REGION Network 319: CARRIER ENCODER POSITION FAULT
   RUNG wire#powerrail
      Contact( "reset" )
      { S7_Templates := "SrcType := Word" } EQ_Contact(in1 := "DB101_DB_SDC_FAULTS".Carrier_Fault[39], in2 := 131)
      Coil( "DB302_HMI_Faults".Carrier39_Faults_0.%X12 )
   END_RUNG
   // the same network as SCL:
   "DB302_HMI_Faults".Carrier39_Faults_0.%X12 := "reset" AND ("DB101_DB_SDC_FAULTS".Carrier_Fault[39] = 131);
END_REGION

REGION Network 320: CARRIER ENCODER INTERNAL ERROR
   RUNG wire#powerrail
      Contact( "reset" )
      { S7_Templates := "SrcType := Word" } EQ_Contact(in1 := "DB101_DB_SDC_FAULTS".Carrier_Fault[39], in2 := 132)
      Coil( "DB302_HMI_Faults".Carrier39_Faults_0.%X13 )
   END_RUNG
   // the same network as SCL:
   "DB302_HMI_Faults".Carrier39_Faults_0.%X13 := "reset" AND ("DB101_DB_SDC_FAULTS".Carrier_Fault[39] = 132);
END_REGION

REGION Network 321: CARRIER ENCODER COMM FAULT
   RUNG wire#powerrail
      Contact( "reset" )
      { S7_Templates := "SrcType := Word" } EQ_Contact(in1 := "DB101_DB_SDC_FAULTS".Carrier_Fault[39], in2 := 133)
      Coil( "DB302_HMI_Faults".Carrier39_Faults_0.%X14 )
   END_RUNG
   // the same network as SCL:
   "DB302_HMI_Faults".Carrier39_Faults_0.%X14 := "reset" AND ("DB101_DB_SDC_FAULTS".Carrier_Fault[39] = 133);
END_REGION

REGION Network 322: CARRIER HMI COMM FAULT
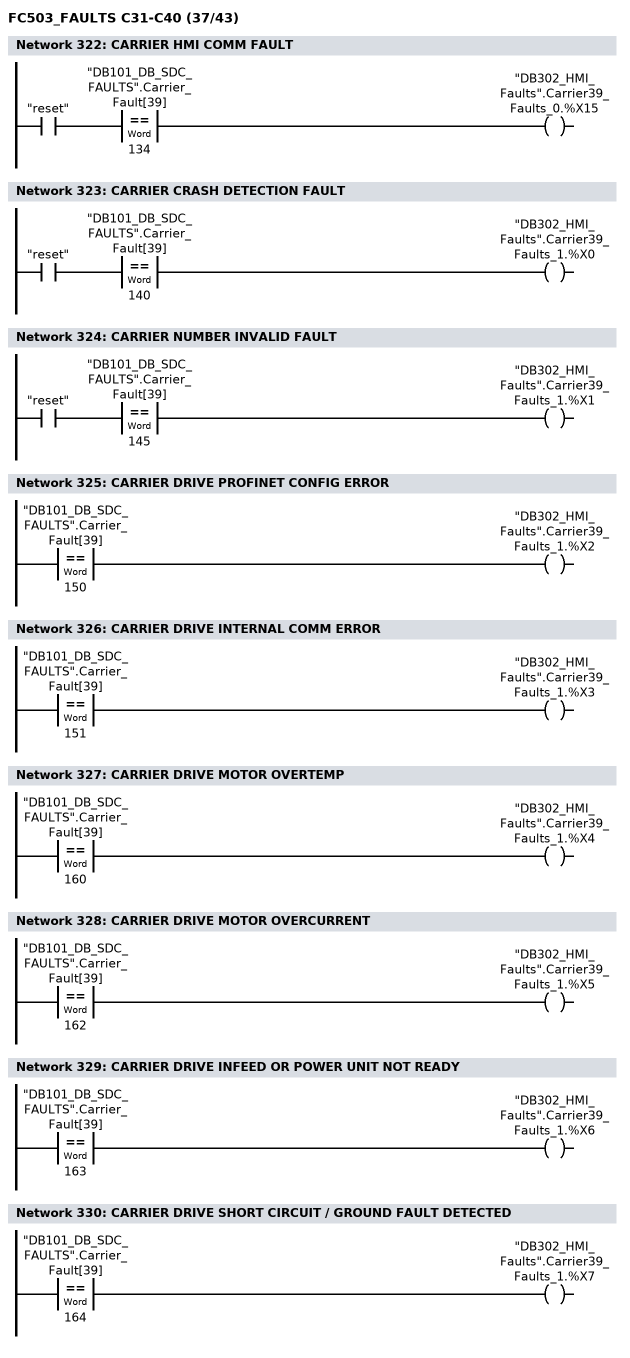
   RUNG wire#powerrail
      Contact( "reset" )
      { S7_Templates := "SrcType := Word" } EQ_Contact(in1 := "DB101_DB_SDC_FAULTS".Carrier_Fault[39], in2 := 134)
      Coil( "DB302_HMI_Faults".Carrier39_Faults_0.%X15 )
   END_RUNG
   // the same network as SCL:
   "DB302_HMI_Faults".Carrier39_Faults_0.%X15 := "reset" AND ("DB101_DB_SDC_FAULTS".Carrier_Fault[39] = 134);
END_REGION

REGION Network 323: CARRIER CRASH DETECTION FAULT
   RUNG wire#powerrail
      Contact( "reset" )
      { S7_Templates := "SrcType := Word" } EQ_Contact(in1 := "DB101_DB_SDC_FAULTS".Carrier_Fault[39], in2 := 140)
      Coil( "DB302_HMI_Faults".Carrier39_Faults_1.%X0 )
   END_RUNG
   // the same network as SCL:
   "DB302_HMI_Faults".Carrier39_Faults_1.%X0 := "reset" AND ("DB101_DB_SDC_FAULTS".Carrier_Fault[39] = 140);
END_REGION

REGION Network 324: CARRIER NUMBER INVALID FAULT
   RUNG wire#powerrail
      Contact( "reset" )
      { S7_Templates := "SrcType := Word" } EQ_Contact(in1 := "DB101_DB_SDC_FAULTS".Carrier_Fault[39], in2 := 145)
      Coil( "DB302_HMI_Faults".Carrier39_Faults_1.%X1 )
   END_RUNG
   // the same network as SCL:
   "DB302_HMI_Faults".Carrier39_Faults_1.%X1 := "reset" AND ("DB101_DB_SDC_FAULTS".Carrier_Fault[39] = 145);
END_REGION

REGION Network 325: CARRIER DRIVE PROFINET CONFIG ERROR
   RUNG wire#powerrail
      { S7_Templates := "SrcType := Word" } EQ_Contact(in1 := "DB101_DB_SDC_FAULTS".Carrier_Fault[39], in2 := 150)
      Coil( "DB302_HMI_Faults".Carrier39_Faults_1.%X2 )
   END_RUNG
   // the same network as SCL:
   "DB302_HMI_Faults".Carrier39_Faults_1.%X2 := "DB101_DB_SDC_FAULTS".Carrier_Fault[39] = 150;
END_REGION

REGION Network 326: CARRIER DRIVE INTERNAL COMM ERROR
   RUNG wire#powerrail
      { S7_Templates := "SrcType := Word" } EQ_Contact(in1 := "DB101_DB_SDC_FAULTS".Carrier_Fault[39], in2 := 151)
      Coil( "DB302_HMI_Faults".Carrier39_Faults_1.%X3 )
   END_RUNG
   // the same network as SCL:
   "DB302_HMI_Faults".Carrier39_Faults_1.%X3 := "DB101_DB_SDC_FAULTS".Carrier_Fault[39] = 151;
END_REGION

REGION Network 327: CARRIER DRIVE MOTOR OVERTEMP
   RUNG wire#powerrail
      { S7_Templates := "SrcType := Word" } EQ_Contact(in1 := "DB101_DB_SDC_FAULTS".Carrier_Fault[39], in2 := 160)
      Coil( "DB302_HMI_Faults".Carrier39_Faults_1.%X4 )
   END_RUNG
   // the same network as SCL:
   "DB302_HMI_Faults".Carrier39_Faults_1.%X4 := "DB101_DB_SDC_FAULTS".Carrier_Fault[39] = 160;
END_REGION

REGION Network 328: CARRIER DRIVE MOTOR OVERCURRENT
   RUNG wire#powerrail
      { S7_Templates := "SrcType := Word" } EQ_Contact(in1 := "DB101_DB_SDC_FAULTS".Carrier_Fault[39], in2 := 162)
      Coil( "DB302_HMI_Faults".Carrier39_Faults_1.%X5 )
   END_RUNG
   // the same network as SCL:
   "DB302_HMI_Faults".Carrier39_Faults_1.%X5 := "DB101_DB_SDC_FAULTS".Carrier_Fault[39] = 162;
END_REGION

REGION Network 329: CARRIER DRIVE INFEED OR POWER UNIT NOT READY
   RUNG wire#powerrail
      { S7_Templates := "SrcType := Word" } EQ_Contact(in1 := "DB101_DB_SDC_FAULTS".Carrier_Fault[39], in2 := 163)
      Coil( "DB302_HMI_Faults".Carrier39_Faults_1.%X6 )
   END_RUNG
   // the same network as SCL:
   "DB302_HMI_Faults".Carrier39_Faults_1.%X6 := "DB101_DB_SDC_FAULTS".Carrier_Fault[39] = 163;
END_REGION

REGION Network 330: CARRIER DRIVE SHORT CIRCUIT / GROUND FAULT DETECTED
   RUNG wire#powerrail
      { S7_Templates := "SrcType := Word" } EQ_Contact(in1 := "DB101_DB_SDC_FAULTS".Carrier_Fault[39], in2 := 164)
      Coil( "DB302_HMI_Faults".Carrier39_Faults_1.%X7 )
   END_RUNG
   // the same network as SCL:
   "DB302_HMI_Faults".Carrier39_Faults_1.%X7 := "DB101_DB_SDC_FAULTS".Carrier_Fault[39] = 164;
END_REGION

REGION Network 331: CARRIER DRIVE PROFINET SETPOINT TIMEOUT
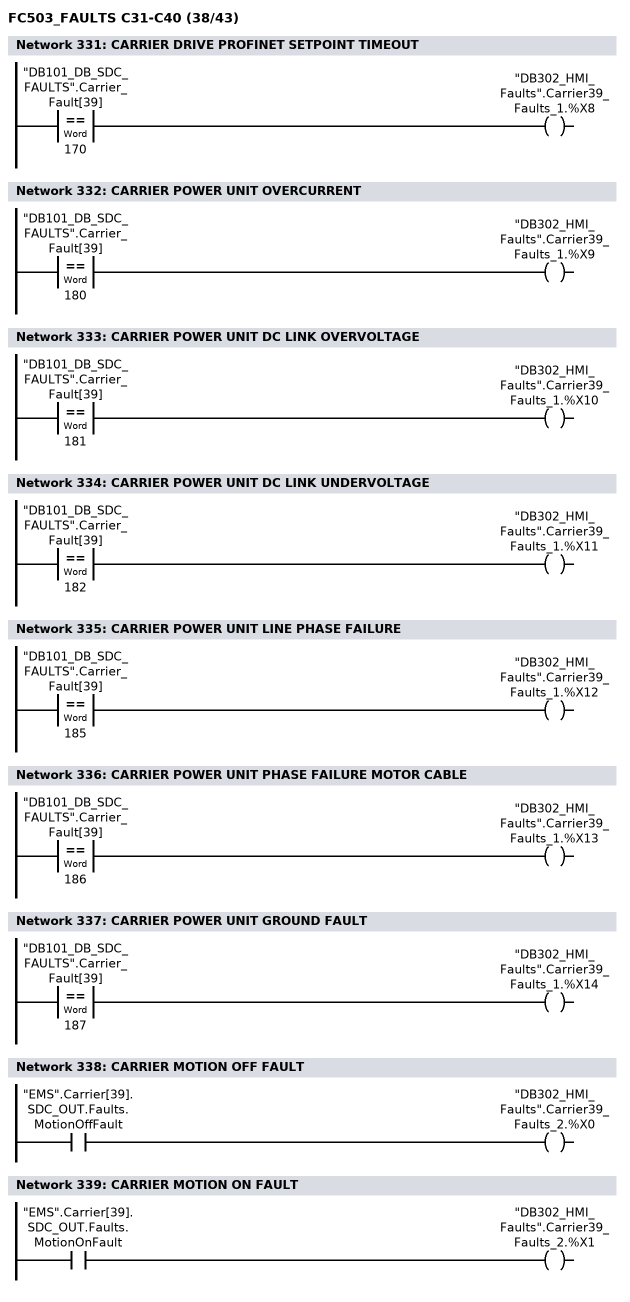
   RUNG wire#powerrail
      { S7_Templates := "SrcType := Word" } EQ_Contact(in1 := "DB101_DB_SDC_FAULTS".Carrier_Fault[39], in2 := 170)
      Coil( "DB302_HMI_Faults".Carrier39_Faults_1.%X8 )
   END_RUNG
   // the same network as SCL:
   "DB302_HMI_Faults".Carrier39_Faults_1.%X8 := "DB101_DB_SDC_FAULTS".Carrier_Fault[39] = 170;
END_REGION

REGION Network 332: CARRIER POWER UNIT OVERCURRENT
   RUNG wire#powerrail
      { S7_Templates := "SrcType := Word" } EQ_Contact(in1 := "DB101_DB_SDC_FAULTS".Carrier_Fault[39], in2 := 180)
      Coil( "DB302_HMI_Faults".Carrier39_Faults_1.%X9 )
   END_RUNG
   // the same network as SCL:
   "DB302_HMI_Faults".Carrier39_Faults_1.%X9 := "DB101_DB_SDC_FAULTS".Carrier_Fault[39] = 180;
END_REGION

REGION Network 333: CARRIER POWER UNIT DC LINK OVERVOLTAGE
   RUNG wire#powerrail
      { S7_Templates := "SrcType := Word" } EQ_Contact(in1 := "DB101_DB_SDC_FAULTS".Carrier_Fault[39], in2 := 181)
      Coil( "DB302_HMI_Faults".Carrier39_Faults_1.%X10 )
   END_RUNG
   // the same network as SCL:
   "DB302_HMI_Faults".Carrier39_Faults_1.%X10 := "DB101_DB_SDC_FAULTS".Carrier_Fault[39] = 181;
END_REGION

REGION Network 334: CARRIER POWER UNIT DC LINK UNDERVOLTAGE
   RUNG wire#powerrail
      { S7_Templates := "SrcType := Word" } EQ_Contact(in1 := "DB101_DB_SDC_FAULTS".Carrier_Fault[39], in2 := 182)
      Coil( "DB302_HMI_Faults".Carrier39_Faults_1.%X11 )
   END_RUNG
   // the same network as SCL:
   "DB302_HMI_Faults".Carrier39_Faults_1.%X11 := "DB101_DB_SDC_FAULTS".Carrier_Fault[39] = 182;
END_REGION

REGION Network 335: CARRIER POWER UNIT LINE PHASE FAILURE
   RUNG wire#powerrail
      { S7_Templates := "SrcType := Word" } EQ_Contact(in1 := "DB101_DB_SDC_FAULTS".Carrier_Fault[39], in2 := 185)
      Coil( "DB302_HMI_Faults".Carrier39_Faults_1.%X12 )
   END_RUNG
   // the same network as SCL:
   "DB302_HMI_Faults".Carrier39_Faults_1.%X12 := "DB101_DB_SDC_FAULTS".Carrier_Fault[39] = 185;
END_REGION

REGION Network 336: CARRIER POWER UNIT PHASE FAILURE MOTOR CABLE
   RUNG wire#powerrail
      { S7_Templates := "SrcType := Word" } EQ_Contact(in1 := "DB101_DB_SDC_FAULTS".Carrier_Fault[39], in2 := 186)
      Coil( "DB302_HMI_Faults".Carrier39_Faults_1.%X13 )
   END_RUNG
   // the same network as SCL:
   "DB302_HMI_Faults".Carrier39_Faults_1.%X13 := "DB101_DB_SDC_FAULTS".Carrier_Fault[39] = 186;
END_REGION

REGION Network 337: CARRIER POWER UNIT GROUND FAULT
   RUNG wire#powerrail
      { S7_Templates := "SrcType := Word" } EQ_Contact(in1 := "DB101_DB_SDC_FAULTS".Carrier_Fault[39], in2 := 187)
      Coil( "DB302_HMI_Faults".Carrier39_Faults_1.%X14 )
   END_RUNG
   // the same network as SCL:
   "DB302_HMI_Faults".Carrier39_Faults_1.%X14 := "DB101_DB_SDC_FAULTS".Carrier_Fault[39] = 187;
END_REGION

REGION Network 338: CARRIER MOTION OFF FAULT
   RUNG wire#powerrail
      Contact( "EMS".Carrier[39].SDC_OUT.Faults.MotionOffFault )
      Coil( "DB302_HMI_Faults".Carrier39_Faults_2.%X0 )
   END_RUNG
   // the same network as SCL:
   "DB302_HMI_Faults".Carrier39_Faults_2.%X0 := "EMS".Carrier[39].SDC_OUT.Faults.MotionOffFault;
END_REGION

REGION Network 339: CARRIER MOTION ON FAULT
   RUNG wire#powerrail
      Contact( "EMS".Carrier[39].SDC_OUT.Faults.MotionOnFault )
      Coil( "DB302_HMI_Faults".Carrier39_Faults_2.%X1 )
   END_RUNG
   // the same network as SCL:
   "DB302_HMI_Faults".Carrier39_Faults_2.%X1 := "EMS".Carrier[39].SDC_OUT.Faults.MotionOnFault;
END_REGION

REGION Network 340: CARRIER SPACING FAULT
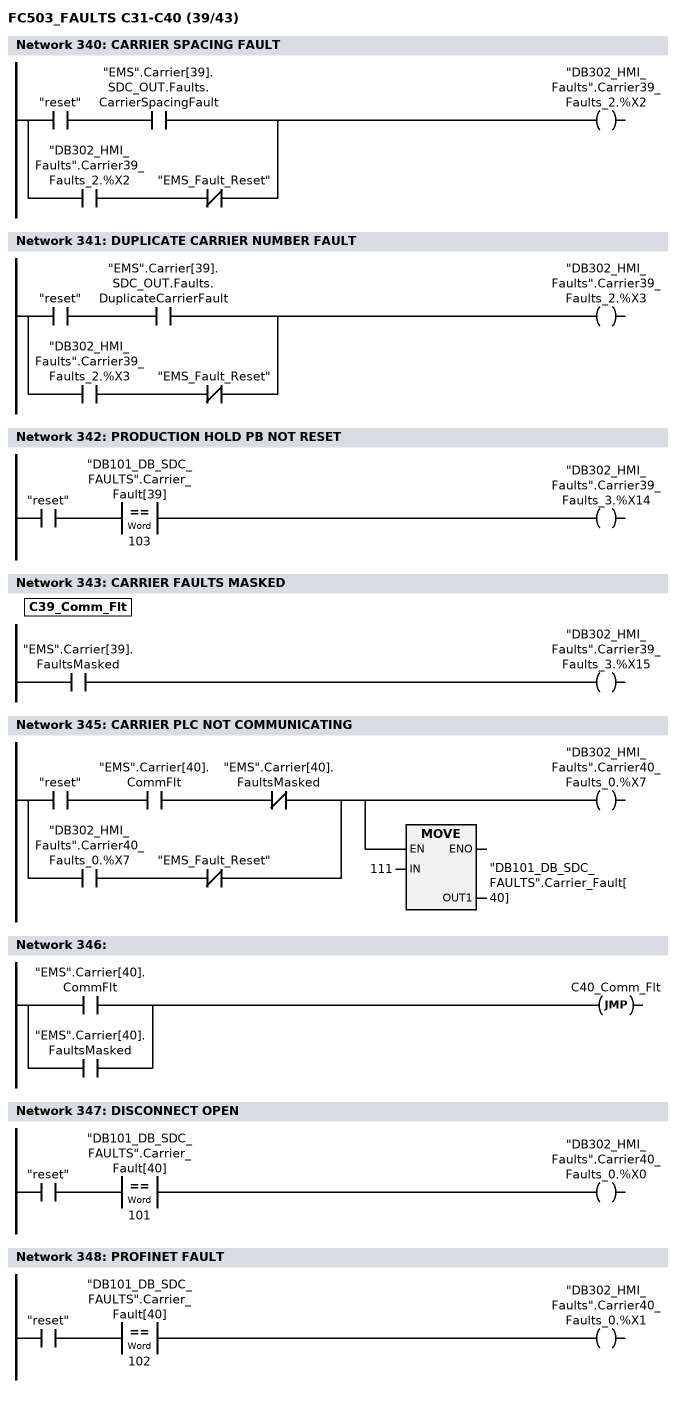
   RUNG wire#powerrail
      Contact( "reset" )
      Contact( "EMS".Carrier[39].SDC_OUT.Faults.CarrierSpacingFault )
      wire#w1
      Coil( "DB302_HMI_Faults".Carrier39_Faults_2.%X2 )
   END_RUNG
   RUNG wire#powerrail
      Contact( "DB302_HMI_Faults".Carrier39_Faults_2.%X2 )
      I_Contact( "EMS_Fault_Reset" )
   END_RUNG wire#w1
   // the same network as SCL:
   "DB302_HMI_Faults".Carrier39_Faults_2.%X2 := ("reset" AND "EMS".Carrier[39].SDC_OUT.Faults.CarrierSpacingFault) OR ("DB302_HMI_Faults".Carrier39_Faults_2.%X2 AND NOT "EMS_Fault_Reset");
END_REGION

REGION Network 341: DUPLICATE CARRIER NUMBER FAULT
   RUNG wire#powerrail
      Contact( "reset" )
      Contact( "EMS".Carrier[39].SDC_OUT.Faults.DuplicateCarrierFault )
      wire#w1
      Coil( "DB302_HMI_Faults".Carrier39_Faults_2.%X3 )
   END_RUNG
   RUNG wire#powerrail
      Contact( "DB302_HMI_Faults".Carrier39_Faults_2.%X3 )
      I_Contact( "EMS_Fault_Reset" )
   END_RUNG wire#w1
   // the same network as SCL:
   "DB302_HMI_Faults".Carrier39_Faults_2.%X3 := ("reset" AND "EMS".Carrier[39].SDC_OUT.Faults.DuplicateCarrierFault) OR ("DB302_HMI_Faults".Carrier39_Faults_2.%X3 AND NOT "EMS_Fault_Reset");
END_REGION

REGION Network 342: PRODUCTION HOLD PB NOT RESET
   RUNG wire#powerrail
      Contact( "reset" )
      { S7_Templates := "SrcType := Word" } EQ_Contact(in1 := "DB101_DB_SDC_FAULTS".Carrier_Fault[39], in2 := 103)
      Coil( "DB302_HMI_Faults".Carrier39_Faults_3.%X14 )
   END_RUNG
   // the same network as SCL:
   "DB302_HMI_Faults".Carrier39_Faults_3.%X14 := "reset" AND ("DB101_DB_SDC_FAULTS".Carrier_Fault[39] = 103);
END_REGION

REGION Network 343: CARRIER FAULTS MASKED
   Label( C39_Comm_Flt )
   RUNG wire#powerrail
      Contact( "EMS".Carrier[39].FaultsMasked )
      Coil( "DB302_HMI_Faults".Carrier39_Faults_3.%X15 )
   END_RUNG
   // the same network as SCL:
   C39_Comm_Flt:
   "DB302_HMI_Faults".Carrier39_Faults_3.%X15 := "EMS".Carrier[39].FaultsMasked;
END_REGION

REGION Network 344: CARRIER 40 FAULTS
END_REGION

REGION Network 345: CARRIER PLC NOT COMMUNICATING
   RUNG wire#powerrail
      Contact( "reset" )
      Contact( "EMS".Carrier[40].CommFlt )
      I_Contact( "EMS".Carrier[40].FaultsMasked )
      wire#w1
      Coil( "DB302_HMI_Faults".Carrier40_Faults_0.%X7 )
   END_RUNG
   RUNG wire#powerrail
      Contact( "DB302_HMI_Faults".Carrier40_Faults_0.%X7 )
      I_Contact( "EMS_Fault_Reset" )
   END_RUNG wire#w1
   RUNG wire#w1
      Move(in := 111, out1 => "DB101_DB_SDC_FAULTS".Carrier_Fault[40])
   END_RUNG
   // the same network as SCL:
   "DB302_HMI_Faults".Carrier40_Faults_0.%X7 := ("reset" AND "EMS".Carrier[40].CommFlt AND NOT "EMS".Carrier[40].FaultsMasked) OR ("DB302_HMI_Faults".Carrier40_Faults_0.%X7 AND NOT "EMS_Fault_Reset");
   IF "DB302_HMI_Faults".Carrier40_Faults_0.%X7 THEN "DB101_DB_SDC_FAULTS".Carrier_Fault[40] := 111; END_IF;
END_REGION

REGION Network 346
   RUNG wire#powerrail
      Contact( "EMS".Carrier[40].CommFlt )
      wire#w1
      JumpCoil( C40_Comm_Flt )
   END_RUNG
   RUNG wire#powerrail
      Contact( "EMS".Carrier[40].FaultsMasked )
   END_RUNG wire#w1
   // the same network as SCL:
   IF "EMS".Carrier[40].CommFlt OR "EMS".Carrier[40].FaultsMasked THEN GOTO C40_Comm_Flt; END_IF;
END_REGION

REGION Network 347: DISCONNECT OPEN
   RUNG wire#powerrail
      Contact( "reset" )
      { S7_Templates := "SrcType := Word" } EQ_Contact(in1 := "DB101_DB_SDC_FAULTS".Carrier_Fault[40], in2 := 101)
      Coil( "DB302_HMI_Faults".Carrier40_Faults_0.%X0 )
   END_RUNG
   // the same network as SCL:
   "DB302_HMI_Faults".Carrier40_Faults_0.%X0 := "reset" AND ("DB101_DB_SDC_FAULTS".Carrier_Fault[40] = 101);
END_REGION

REGION Network 348: PROFINET FAULT
   RUNG wire#powerrail
      Contact( "reset" )
      { S7_Templates := "SrcType := Word" } EQ_Contact(in1 := "DB101_DB_SDC_FAULTS".Carrier_Fault[40], in2 := 102)
      Coil( "DB302_HMI_Faults".Carrier40_Faults_0.%X1 )
   END_RUNG
   // the same network as SCL:
   "DB302_HMI_Faults".Carrier40_Faults_0.%X1 := "reset" AND ("DB101_DB_SDC_FAULTS".Carrier_Fault[40] = 102);
END_REGION

REGION Network 349: CB2122 TRIPPED
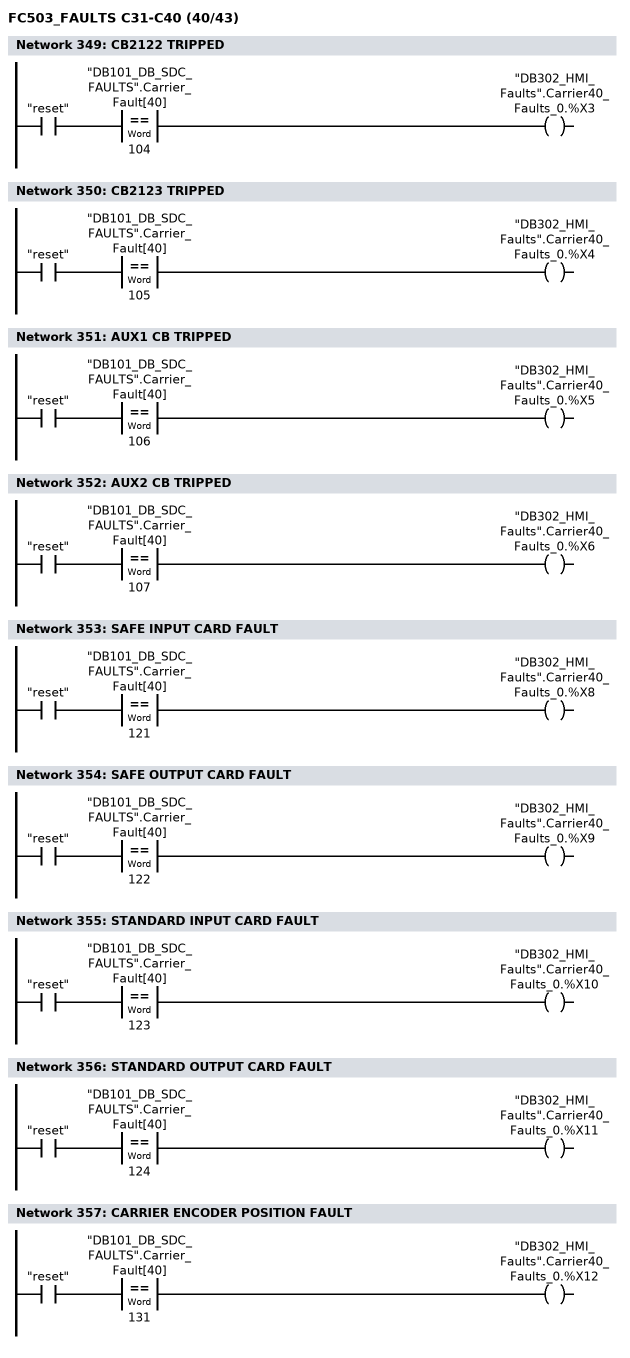
   RUNG wire#powerrail
      Contact( "reset" )
      { S7_Templates := "SrcType := Word" } EQ_Contact(in1 := "DB101_DB_SDC_FAULTS".Carrier_Fault[40], in2 := 104)
      Coil( "DB302_HMI_Faults".Carrier40_Faults_0.%X3 )
   END_RUNG
   // the same network as SCL:
   "DB302_HMI_Faults".Carrier40_Faults_0.%X3 := "reset" AND ("DB101_DB_SDC_FAULTS".Carrier_Fault[40] = 104);
END_REGION

REGION Network 350: CB2123 TRIPPED
   RUNG wire#powerrail
      Contact( "reset" )
      { S7_Templates := "SrcType := Word" } EQ_Contact(in1 := "DB101_DB_SDC_FAULTS".Carrier_Fault[40], in2 := 105)
      Coil( "DB302_HMI_Faults".Carrier40_Faults_0.%X4 )
   END_RUNG
   // the same network as SCL:
   "DB302_HMI_Faults".Carrier40_Faults_0.%X4 := "reset" AND ("DB101_DB_SDC_FAULTS".Carrier_Fault[40] = 105);
END_REGION

REGION Network 351: AUX1 CB TRIPPED
   RUNG wire#powerrail
      Contact( "reset" )
      { S7_Templates := "SrcType := Word" } EQ_Contact(in1 := "DB101_DB_SDC_FAULTS".Carrier_Fault[40], in2 := 106)
      Coil( "DB302_HMI_Faults".Carrier40_Faults_0.%X5 )
   END_RUNG
   // the same network as SCL:
   "DB302_HMI_Faults".Carrier40_Faults_0.%X5 := "reset" AND ("DB101_DB_SDC_FAULTS".Carrier_Fault[40] = 106);
END_REGION

REGION Network 352: AUX2 CB TRIPPED
   RUNG wire#powerrail
      Contact( "reset" )
      { S7_Templates := "SrcType := Word" } EQ_Contact(in1 := "DB101_DB_SDC_FAULTS".Carrier_Fault[40], in2 := 107)
      Coil( "DB302_HMI_Faults".Carrier40_Faults_0.%X6 )
   END_RUNG
   // the same network as SCL:
   "DB302_HMI_Faults".Carrier40_Faults_0.%X6 := "reset" AND ("DB101_DB_SDC_FAULTS".Carrier_Fault[40] = 107);
END_REGION

REGION Network 353: SAFE INPUT CARD FAULT
   RUNG wire#powerrail
      Contact( "reset" )
      { S7_Templates := "SrcType := Word" } EQ_Contact(in1 := "DB101_DB_SDC_FAULTS".Carrier_Fault[40], in2 := 121)
      Coil( "DB302_HMI_Faults".Carrier40_Faults_0.%X8 )
   END_RUNG
   // the same network as SCL:
   "DB302_HMI_Faults".Carrier40_Faults_0.%X8 := "reset" AND ("DB101_DB_SDC_FAULTS".Carrier_Fault[40] = 121);
END_REGION

REGION Network 354: SAFE OUTPUT CARD FAULT
   RUNG wire#powerrail
      Contact( "reset" )
      { S7_Templates := "SrcType := Word" } EQ_Contact(in1 := "DB101_DB_SDC_FAULTS".Carrier_Fault[40], in2 := 122)
      Coil( "DB302_HMI_Faults".Carrier40_Faults_0.%X9 )
   END_RUNG
   // the same network as SCL:
   "DB302_HMI_Faults".Carrier40_Faults_0.%X9 := "reset" AND ("DB101_DB_SDC_FAULTS".Carrier_Fault[40] = 122);
END_REGION

REGION Network 355: STANDARD INPUT CARD FAULT
   RUNG wire#powerrail
      Contact( "reset" )
      { S7_Templates := "SrcType := Word" } EQ_Contact(in1 := "DB101_DB_SDC_FAULTS".Carrier_Fault[40], in2 := 123)
      Coil( "DB302_HMI_Faults".Carrier40_Faults_0.%X10 )
   END_RUNG
   // the same network as SCL:
   "DB302_HMI_Faults".Carrier40_Faults_0.%X10 := "reset" AND ("DB101_DB_SDC_FAULTS".Carrier_Fault[40] = 123);
END_REGION

REGION Network 356: STANDARD OUTPUT CARD FAULT
   RUNG wire#powerrail
      Contact( "reset" )
      { S7_Templates := "SrcType := Word" } EQ_Contact(in1 := "DB101_DB_SDC_FAULTS".Carrier_Fault[40], in2 := 124)
      Coil( "DB302_HMI_Faults".Carrier40_Faults_0.%X11 )
   END_RUNG
   // the same network as SCL:
   "DB302_HMI_Faults".Carrier40_Faults_0.%X11 := "reset" AND ("DB101_DB_SDC_FAULTS".Carrier_Fault[40] = 124);
END_REGION

REGION Network 357: CARRIER ENCODER POSITION FAULT
   RUNG wire#powerrail
      Contact( "reset" )
      { S7_Templates := "SrcType := Word" } EQ_Contact(in1 := "DB101_DB_SDC_FAULTS".Carrier_Fault[40], in2 := 131)
      Coil( "DB302_HMI_Faults".Carrier40_Faults_0.%X12 )
   END_RUNG
   // the same network as SCL:
   "DB302_HMI_Faults".Carrier40_Faults_0.%X12 := "reset" AND ("DB101_DB_SDC_FAULTS".Carrier_Fault[40] = 131);
END_REGION

REGION Network 358: CARRIER ENCODER INTERNAL ERROR
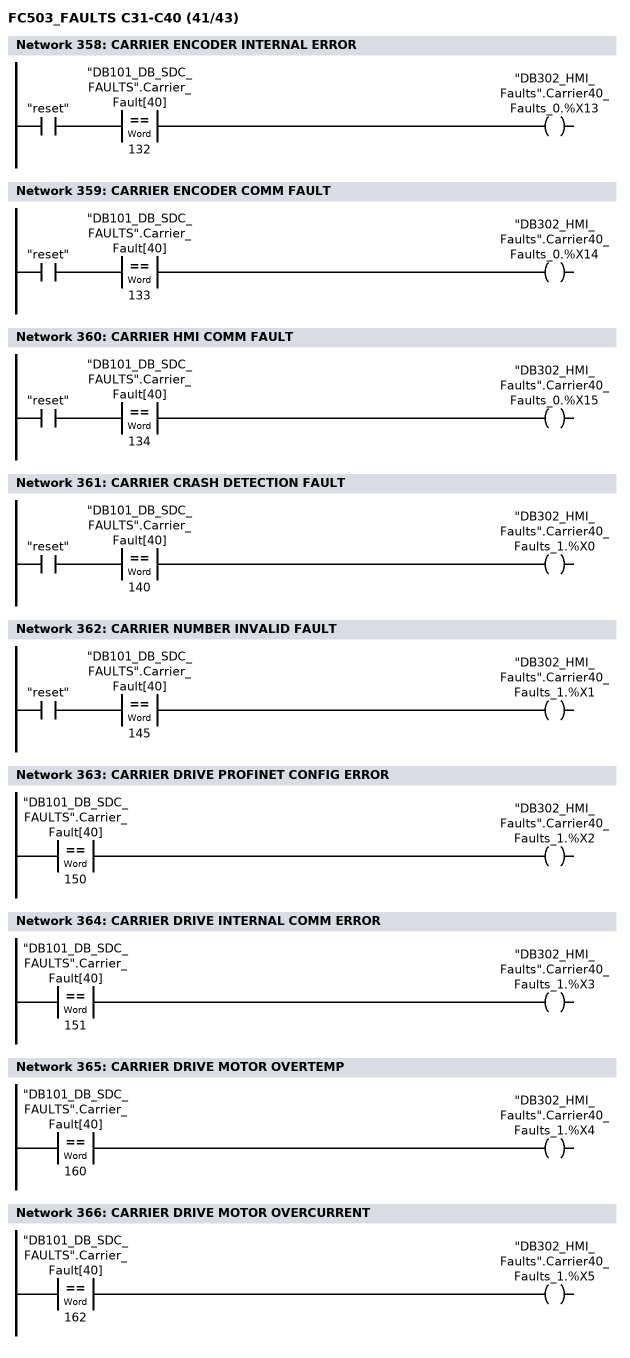
   RUNG wire#powerrail
      Contact( "reset" )
      { S7_Templates := "SrcType := Word" } EQ_Contact(in1 := "DB101_DB_SDC_FAULTS".Carrier_Fault[40], in2 := 132)
      Coil( "DB302_HMI_Faults".Carrier40_Faults_0.%X13 )
   END_RUNG
   // the same network as SCL:
   "DB302_HMI_Faults".Carrier40_Faults_0.%X13 := "reset" AND ("DB101_DB_SDC_FAULTS".Carrier_Fault[40] = 132);
END_REGION

REGION Network 359: CARRIER ENCODER COMM FAULT
   RUNG wire#powerrail
      Contact( "reset" )
      { S7_Templates := "SrcType := Word" } EQ_Contact(in1 := "DB101_DB_SDC_FAULTS".Carrier_Fault[40], in2 := 133)
      Coil( "DB302_HMI_Faults".Carrier40_Faults_0.%X14 )
   END_RUNG
   // the same network as SCL:
   "DB302_HMI_Faults".Carrier40_Faults_0.%X14 := "reset" AND ("DB101_DB_SDC_FAULTS".Carrier_Fault[40] = 133);
END_REGION

REGION Network 360: CARRIER HMI COMM FAULT
   RUNG wire#powerrail
      Contact( "reset" )
      { S7_Templates := "SrcType := Word" } EQ_Contact(in1 := "DB101_DB_SDC_FAULTS".Carrier_Fault[40], in2 := 134)
      Coil( "DB302_HMI_Faults".Carrier40_Faults_0.%X15 )
   END_RUNG
   // the same network as SCL:
   "DB302_HMI_Faults".Carrier40_Faults_0.%X15 := "reset" AND ("DB101_DB_SDC_FAULTS".Carrier_Fault[40] = 134);
END_REGION

REGION Network 361: CARRIER CRASH DETECTION FAULT
   RUNG wire#powerrail
      Contact( "reset" )
      { S7_Templates := "SrcType := Word" } EQ_Contact(in1 := "DB101_DB_SDC_FAULTS".Carrier_Fault[40], in2 := 140)
      Coil( "DB302_HMI_Faults".Carrier40_Faults_1.%X0 )
   END_RUNG
   // the same network as SCL:
   "DB302_HMI_Faults".Carrier40_Faults_1.%X0 := "reset" AND ("DB101_DB_SDC_FAULTS".Carrier_Fault[40] = 140);
END_REGION

REGION Network 362: CARRIER NUMBER INVALID FAULT
   RUNG wire#powerrail
      Contact( "reset" )
      { S7_Templates := "SrcType := Word" } EQ_Contact(in1 := "DB101_DB_SDC_FAULTS".Carrier_Fault[40], in2 := 145)
      Coil( "DB302_HMI_Faults".Carrier40_Faults_1.%X1 )
   END_RUNG
   // the same network as SCL:
   "DB302_HMI_Faults".Carrier40_Faults_1.%X1 := "reset" AND ("DB101_DB_SDC_FAULTS".Carrier_Fault[40] = 145);
END_REGION

REGION Network 363: CARRIER DRIVE PROFINET CONFIG ERROR
   RUNG wire#powerrail
      { S7_Templates := "SrcType := Word" } EQ_Contact(in1 := "DB101_DB_SDC_FAULTS".Carrier_Fault[40], in2 := 150)
      Coil( "DB302_HMI_Faults".Carrier40_Faults_1.%X2 )
   END_RUNG
   // the same network as SCL:
   "DB302_HMI_Faults".Carrier40_Faults_1.%X2 := "DB101_DB_SDC_FAULTS".Carrier_Fault[40] = 150;
END_REGION

REGION Network 364: CARRIER DRIVE INTERNAL COMM ERROR
   RUNG wire#powerrail
      { S7_Templates := "SrcType := Word" } EQ_Contact(in1 := "DB101_DB_SDC_FAULTS".Carrier_Fault[40], in2 := 151)
      Coil( "DB302_HMI_Faults".Carrier40_Faults_1.%X3 )
   END_RUNG
   // the same network as SCL:
   "DB302_HMI_Faults".Carrier40_Faults_1.%X3 := "DB101_DB_SDC_FAULTS".Carrier_Fault[40] = 151;
END_REGION

REGION Network 365: CARRIER DRIVE MOTOR OVERTEMP
   RUNG wire#powerrail
      { S7_Templates := "SrcType := Word" } EQ_Contact(in1 := "DB101_DB_SDC_FAULTS".Carrier_Fault[40], in2 := 160)
      Coil( "DB302_HMI_Faults".Carrier40_Faults_1.%X4 )
   END_RUNG
   // the same network as SCL:
   "DB302_HMI_Faults".Carrier40_Faults_1.%X4 := "DB101_DB_SDC_FAULTS".Carrier_Fault[40] = 160;
END_REGION

REGION Network 366: CARRIER DRIVE MOTOR OVERCURRENT
   RUNG wire#powerrail
      { S7_Templates := "SrcType := Word" } EQ_Contact(in1 := "DB101_DB_SDC_FAULTS".Carrier_Fault[40], in2 := 162)
      Coil( "DB302_HMI_Faults".Carrier40_Faults_1.%X5 )
   END_RUNG
   // the same network as SCL:
   "DB302_HMI_Faults".Carrier40_Faults_1.%X5 := "DB101_DB_SDC_FAULTS".Carrier_Fault[40] = 162;
END_REGION

REGION Network 367: CARRIER DRIVE INFEED OR POWER UNIT NOT READY
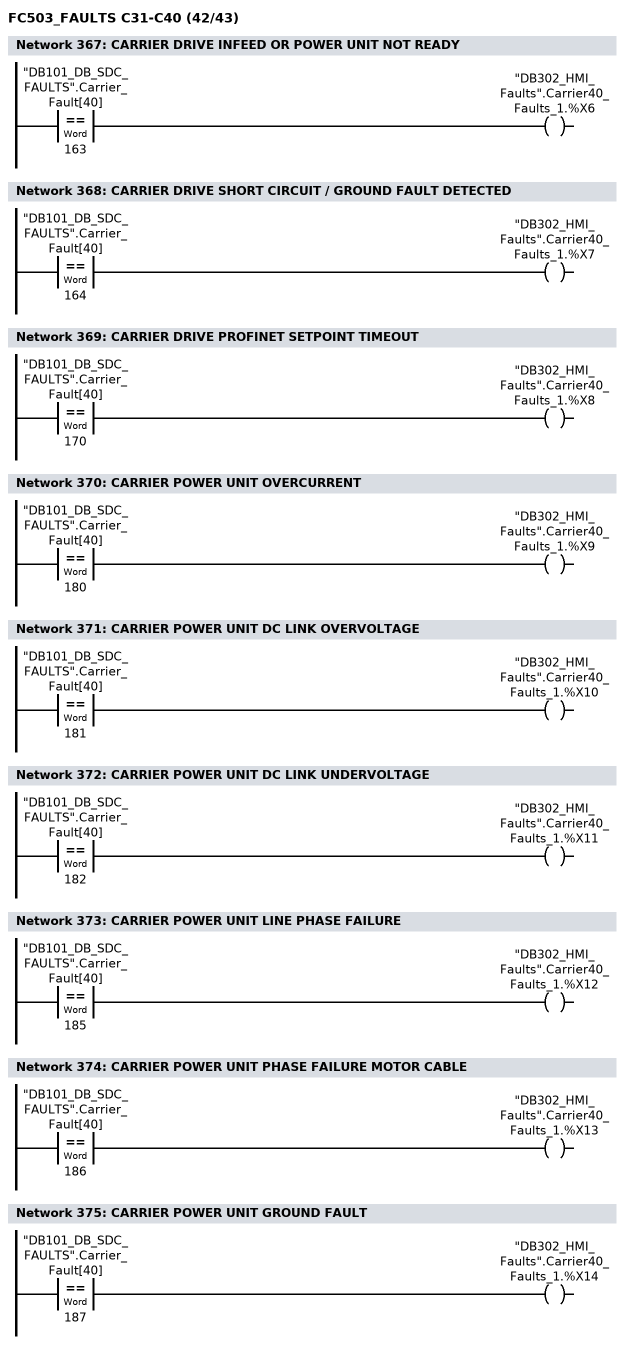
   RUNG wire#powerrail
      { S7_Templates := "SrcType := Word" } EQ_Contact(in1 := "DB101_DB_SDC_FAULTS".Carrier_Fault[40], in2 := 163)
      Coil( "DB302_HMI_Faults".Carrier40_Faults_1.%X6 )
   END_RUNG
   // the same network as SCL:
   "DB302_HMI_Faults".Carrier40_Faults_1.%X6 := "DB101_DB_SDC_FAULTS".Carrier_Fault[40] = 163;
END_REGION

REGION Network 368: CARRIER DRIVE SHORT CIRCUIT / GROUND FAULT DETECTED
   RUNG wire#powerrail
      { S7_Templates := "SrcType := Word" } EQ_Contact(in1 := "DB101_DB_SDC_FAULTS".Carrier_Fault[40], in2 := 164)
      Coil( "DB302_HMI_Faults".Carrier40_Faults_1.%X7 )
   END_RUNG
   // the same network as SCL:
   "DB302_HMI_Faults".Carrier40_Faults_1.%X7 := "DB101_DB_SDC_FAULTS".Carrier_Fault[40] = 164;
END_REGION

REGION Network 369: CARRIER DRIVE PROFINET SETPOINT TIMEOUT
   RUNG wire#powerrail
      { S7_Templates := "SrcType := Word" } EQ_Contact(in1 := "DB101_DB_SDC_FAULTS".Carrier_Fault[40], in2 := 170)
      Coil( "DB302_HMI_Faults".Carrier40_Faults_1.%X8 )
   END_RUNG
   // the same network as SCL:
   "DB302_HMI_Faults".Carrier40_Faults_1.%X8 := "DB101_DB_SDC_FAULTS".Carrier_Fault[40] = 170;
END_REGION

REGION Network 370: CARRIER POWER UNIT OVERCURRENT
   RUNG wire#powerrail
      { S7_Templates := "SrcType := Word" } EQ_Contact(in1 := "DB101_DB_SDC_FAULTS".Carrier_Fault[40], in2 := 180)
      Coil( "DB302_HMI_Faults".Carrier40_Faults_1.%X9 )
   END_RUNG
   // the same network as SCL:
   "DB302_HMI_Faults".Carrier40_Faults_1.%X9 := "DB101_DB_SDC_FAULTS".Carrier_Fault[40] = 180;
END_REGION

REGION Network 371: CARRIER POWER UNIT DC LINK OVERVOLTAGE
   RUNG wire#powerrail
      { S7_Templates := "SrcType := Word" } EQ_Contact(in1 := "DB101_DB_SDC_FAULTS".Carrier_Fault[40], in2 := 181)
      Coil( "DB302_HMI_Faults".Carrier40_Faults_1.%X10 )
   END_RUNG
   // the same network as SCL:
   "DB302_HMI_Faults".Carrier40_Faults_1.%X10 := "DB101_DB_SDC_FAULTS".Carrier_Fault[40] = 181;
END_REGION

REGION Network 372: CARRIER POWER UNIT DC LINK UNDERVOLTAGE
   RUNG wire#powerrail
      { S7_Templates := "SrcType := Word" } EQ_Contact(in1 := "DB101_DB_SDC_FAULTS".Carrier_Fault[40], in2 := 182)
      Coil( "DB302_HMI_Faults".Carrier40_Faults_1.%X11 )
   END_RUNG
   // the same network as SCL:
   "DB302_HMI_Faults".Carrier40_Faults_1.%X11 := "DB101_DB_SDC_FAULTS".Carrier_Fault[40] = 182;
END_REGION

REGION Network 373: CARRIER POWER UNIT LINE PHASE FAILURE
   RUNG wire#powerrail
      { S7_Templates := "SrcType := Word" } EQ_Contact(in1 := "DB101_DB_SDC_FAULTS".Carrier_Fault[40], in2 := 185)
      Coil( "DB302_HMI_Faults".Carrier40_Faults_1.%X12 )
   END_RUNG
   // the same network as SCL:
   "DB302_HMI_Faults".Carrier40_Faults_1.%X12 := "DB101_DB_SDC_FAULTS".Carrier_Fault[40] = 185;
END_REGION

REGION Network 374: CARRIER POWER UNIT PHASE FAILURE MOTOR CABLE
   RUNG wire#powerrail
      { S7_Templates := "SrcType := Word" } EQ_Contact(in1 := "DB101_DB_SDC_FAULTS".Carrier_Fault[40], in2 := 186)
      Coil( "DB302_HMI_Faults".Carrier40_Faults_1.%X13 )
   END_RUNG
   // the same network as SCL:
   "DB302_HMI_Faults".Carrier40_Faults_1.%X13 := "DB101_DB_SDC_FAULTS".Carrier_Fault[40] = 186;
END_REGION

REGION Network 375: CARRIER POWER UNIT GROUND FAULT
   RUNG wire#powerrail
      { S7_Templates := "SrcType := Word" } EQ_Contact(in1 := "DB101_DB_SDC_FAULTS".Carrier_Fault[40], in2 := 187)
      Coil( "DB302_HMI_Faults".Carrier40_Faults_1.%X14 )
   END_RUNG
   // the same network as SCL:
   "DB302_HMI_Faults".Carrier40_Faults_1.%X14 := "DB101_DB_SDC_FAULTS".Carrier_Fault[40] = 187;
END_REGION

REGION Network 376: CARRIER MOTION OFF FAULT
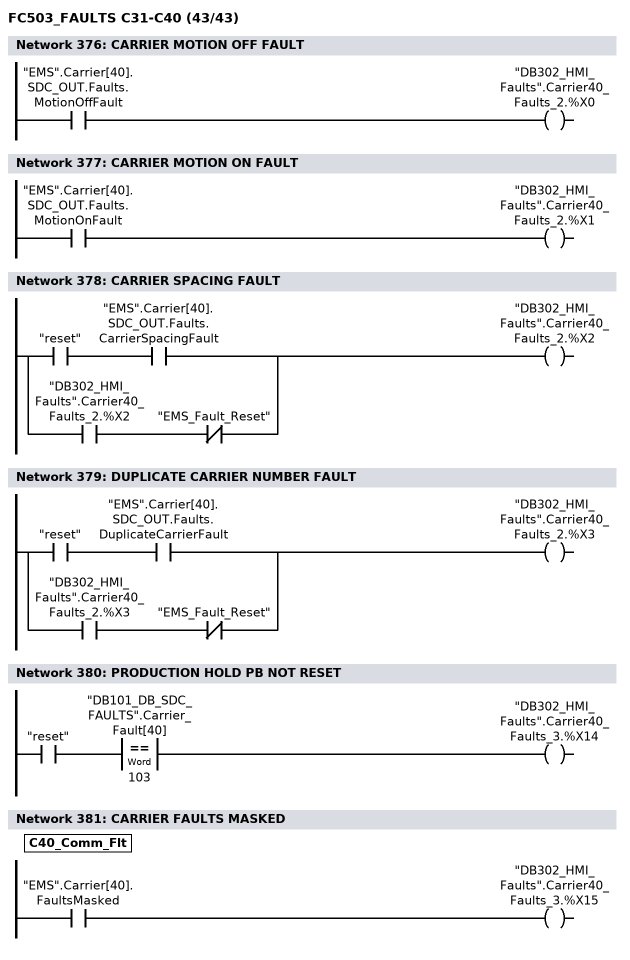
   RUNG wire#powerrail
      Contact( "EMS".Carrier[40].SDC_OUT.Faults.MotionOffFault )
      Coil( "DB302_HMI_Faults".Carrier40_Faults_2.%X0 )
   END_RUNG
   // the same network as SCL:
   "DB302_HMI_Faults".Carrier40_Faults_2.%X0 := "EMS".Carrier[40].SDC_OUT.Faults.MotionOffFault;
END_REGION

REGION Network 377: CARRIER MOTION ON FAULT
   RUNG wire#powerrail
      Contact( "EMS".Carrier[40].SDC_OUT.Faults.MotionOnFault )
      Coil( "DB302_HMI_Faults".Carrier40_Faults_2.%X1 )
   END_RUNG
   // the same network as SCL:
   "DB302_HMI_Faults".Carrier40_Faults_2.%X1 := "EMS".Carrier[40].SDC_OUT.Faults.MotionOnFault;
END_REGION

REGION Network 378: CARRIER SPACING FAULT
   RUNG wire#powerrail
      Contact( "reset" )
      Contact( "EMS".Carrier[40].SDC_OUT.Faults.CarrierSpacingFault )
      wire#w1
      Coil( "DB302_HMI_Faults".Carrier40_Faults_2.%X2 )
   END_RUNG
   RUNG wire#powerrail
      Contact( "DB302_HMI_Faults".Carrier40_Faults_2.%X2 )
      I_Contact( "EMS_Fault_Reset" )
   END_RUNG wire#w1
   // the same network as SCL:
   "DB302_HMI_Faults".Carrier40_Faults_2.%X2 := ("reset" AND "EMS".Carrier[40].SDC_OUT.Faults.CarrierSpacingFault) OR ("DB302_HMI_Faults".Carrier40_Faults_2.%X2 AND NOT "EMS_Fault_Reset");
END_REGION

REGION Network 379: DUPLICATE CARRIER NUMBER FAULT
   RUNG wire#powerrail
      Contact( "reset" )
      Contact( "EMS".Carrier[40].SDC_OUT.Faults.DuplicateCarrierFault )
      wire#w1
      Coil( "DB302_HMI_Faults".Carrier40_Faults_2.%X3 )
   END_RUNG
   RUNG wire#powerrail
      Contact( "DB302_HMI_Faults".Carrier40_Faults_2.%X3 )
      I_Contact( "EMS_Fault_Reset" )
   END_RUNG wire#w1
   // the same network as SCL:
   "DB302_HMI_Faults".Carrier40_Faults_2.%X3 := ("reset" AND "EMS".Carrier[40].SDC_OUT.Faults.DuplicateCarrierFault) OR ("DB302_HMI_Faults".Carrier40_Faults_2.%X3 AND NOT "EMS_Fault_Reset");
END_REGION

REGION Network 380: PRODUCTION HOLD PB NOT RESET
   RUNG wire#powerrail
      Contact( "reset" )
      { S7_Templates := "SrcType := Word" } EQ_Contact(in1 := "DB101_DB_SDC_FAULTS".Carrier_Fault[40], in2 := 103)
      Coil( "DB302_HMI_Faults".Carrier40_Faults_3.%X14 )
   END_RUNG
   // the same network as SCL:
   "DB302_HMI_Faults".Carrier40_Faults_3.%X14 := "reset" AND ("DB101_DB_SDC_FAULTS".Carrier_Fault[40] = 103);
END_REGION

REGION Network 381: CARRIER FAULTS MASKED
   Label( C40_Comm_Flt )
   RUNG wire#powerrail
      Contact( "EMS".Carrier[40].FaultsMasked )
      Coil( "DB302_HMI_Faults".Carrier40_Faults_3.%X15 )
   END_RUNG
   // the same network as SCL:
   C40_Comm_Flt:
   "DB302_HMI_Faults".Carrier40_Faults_3.%X15 := "EMS".Carrier[40].FaultsMasked;
END_REGION
END_FUNCTION

FUNCTION "FC504_FAULTS C41-C50" : Void   // FC504, LAD
{ S7_Optimized_Access := 'TRUE' }
VERSION : 0.1
BEGIN

REGION Network 1: CARRIER 41 FAULTS
END_REGION

REGION Network 2: CARRIER PLC NOT COMMUNICATING
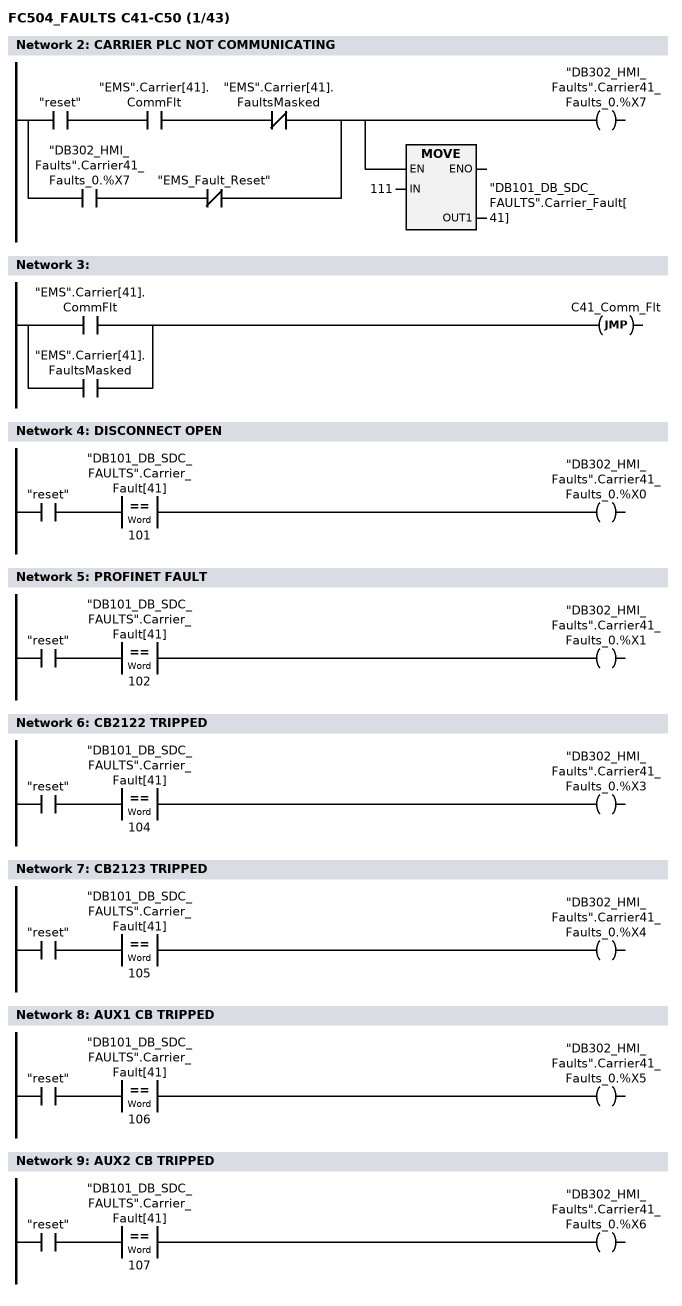
   RUNG wire#powerrail
      Contact( "reset" )
      Contact( "EMS".Carrier[41].CommFlt )
      I_Contact( "EMS".Carrier[41].FaultsMasked )
      wire#w1
      Coil( "DB302_HMI_Faults".Carrier41_Faults_0.%X7 )
   END_RUNG
   RUNG wire#powerrail
      Contact( "DB302_HMI_Faults".Carrier41_Faults_0.%X7 )
      I_Contact( "EMS_Fault_Reset" )
   END_RUNG wire#w1
   RUNG wire#w1
      Move(in := 111, out1 => "DB101_DB_SDC_FAULTS".Carrier_Fault[41])
   END_RUNG
   // the same network as SCL:
   "DB302_HMI_Faults".Carrier41_Faults_0.%X7 := ("reset" AND "EMS".Carrier[41].CommFlt AND NOT "EMS".Carrier[41].FaultsMasked) OR ("DB302_HMI_Faults".Carrier41_Faults_0.%X7 AND NOT "EMS_Fault_Reset");
   IF "DB302_HMI_Faults".Carrier41_Faults_0.%X7 THEN "DB101_DB_SDC_FAULTS".Carrier_Fault[41] := 111; END_IF;
END_REGION

REGION Network 3
   RUNG wire#powerrail
      Contact( "EMS".Carrier[41].CommFlt )
      wire#w1
      JumpCoil( C41_Comm_Flt )
   END_RUNG
   RUNG wire#powerrail
      Contact( "EMS".Carrier[41].FaultsMasked )
   END_RUNG wire#w1
   // the same network as SCL:
   IF "EMS".Carrier[41].CommFlt OR "EMS".Carrier[41].FaultsMasked THEN GOTO C41_Comm_Flt; END_IF;
END_REGION

REGION Network 4: DISCONNECT OPEN
   RUNG wire#powerrail
      Contact( "reset" )
      { S7_Templates := "SrcType := Word" } EQ_Contact(in1 := "DB101_DB_SDC_FAULTS".Carrier_Fault[41], in2 := 101)
      Coil( "DB302_HMI_Faults".Carrier41_Faults_0.%X0 )
   END_RUNG
   // the same network as SCL:
   "DB302_HMI_Faults".Carrier41_Faults_0.%X0 := "reset" AND ("DB101_DB_SDC_FAULTS".Carrier_Fault[41] = 101);
END_REGION

REGION Network 5: PROFINET FAULT
   RUNG wire#powerrail
      Contact( "reset" )
      { S7_Templates := "SrcType := Word" } EQ_Contact(in1 := "DB101_DB_SDC_FAULTS".Carrier_Fault[41], in2 := 102)
      Coil( "DB302_HMI_Faults".Carrier41_Faults_0.%X1 )
   END_RUNG
   // the same network as SCL:
   "DB302_HMI_Faults".Carrier41_Faults_0.%X1 := "reset" AND ("DB101_DB_SDC_FAULTS".Carrier_Fault[41] = 102);
END_REGION

REGION Network 6: CB2122 TRIPPED
   RUNG wire#powerrail
      Contact( "reset" )
      { S7_Templates := "SrcType := Word" } EQ_Contact(in1 := "DB101_DB_SDC_FAULTS".Carrier_Fault[41], in2 := 104)
      Coil( "DB302_HMI_Faults".Carrier41_Faults_0.%X3 )
   END_RUNG
   // the same network as SCL:
   "DB302_HMI_Faults".Carrier41_Faults_0.%X3 := "reset" AND ("DB101_DB_SDC_FAULTS".Carrier_Fault[41] = 104);
END_REGION

REGION Network 7: CB2123 TRIPPED
   RUNG wire#powerrail
      Contact( "reset" )
      { S7_Templates := "SrcType := Word" } EQ_Contact(in1 := "DB101_DB_SDC_FAULTS".Carrier_Fault[41], in2 := 105)
      Coil( "DB302_HMI_Faults".Carrier41_Faults_0.%X4 )
   END_RUNG
   // the same network as SCL:
   "DB302_HMI_Faults".Carrier41_Faults_0.%X4 := "reset" AND ("DB101_DB_SDC_FAULTS".Carrier_Fault[41] = 105);
END_REGION

REGION Network 8: AUX1 CB TRIPPED
   RUNG wire#powerrail
      Contact( "reset" )
      { S7_Templates := "SrcType := Word" } EQ_Contact(in1 := "DB101_DB_SDC_FAULTS".Carrier_Fault[41], in2 := 106)
      Coil( "DB302_HMI_Faults".Carrier41_Faults_0.%X5 )
   END_RUNG
   // the same network as SCL:
   "DB302_HMI_Faults".Carrier41_Faults_0.%X5 := "reset" AND ("DB101_DB_SDC_FAULTS".Carrier_Fault[41] = 106);
END_REGION

REGION Network 9: AUX2 CB TRIPPED
   RUNG wire#powerrail
      Contact( "reset" )
      { S7_Templates := "SrcType := Word" } EQ_Contact(in1 := "DB101_DB_SDC_FAULTS".Carrier_Fault[41], in2 := 107)
      Coil( "DB302_HMI_Faults".Carrier41_Faults_0.%X6 )
   END_RUNG
   // the same network as SCL:
   "DB302_HMI_Faults".Carrier41_Faults_0.%X6 := "reset" AND ("DB101_DB_SDC_FAULTS".Carrier_Fault[41] = 107);
END_REGION

REGION Network 10: SAFE INPUT CARD FAULT
